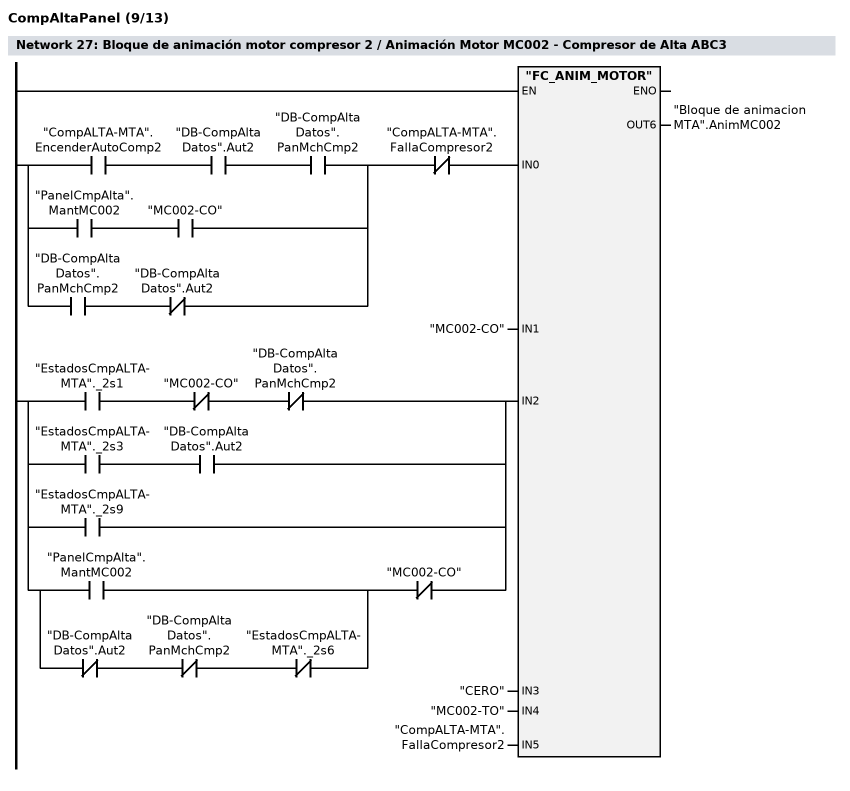
   RUNG wire#powerrail
      "FC_ANIM_MOTOR"(IN0 := wire#w2, IN2 := wire#w4, IN1 := "MC002-CO", IN3 := "CERO", IN4 := "MC002-TO", IN5 := "CompALTA-MTA".FallaCompresor2, OUT6 => "Bloque de animacion MTA".AnimMC002)
   END_RUNG
   RUNG wire#powerrail
      Contact( "CompALTA-MTA".EncenderAutoComp2 )
      Contact( "DB-CompAltaDatos".Aut2 )
      Contact( "DB-CompAltaDatos".PanMchCmp2 )
      wire#w1
      I_Contact( "CompALTA-MTA".FallaCompresor2 )
   END_RUNG wire#w2
   RUNG wire#powerrail
      Contact( "PanelCmpAlta".MantMC002 )
      Contact( "MC002-CO" )
   END_RUNG wire#w1
   RUNG wire#powerrail
      Contact( "DB-CompAltaDatos".PanMchCmp2 )
      I_Contact( "DB-CompAltaDatos".Aut2 )
   END_RUNG wire#w1
   RUNG wire#powerrail
      Contact( "EstadosCmpALTA-MTA"._2s1 )
      I_Contact( "MC002-CO" )
      I_Contact( "DB-CompAltaDatos".PanMchCmp2 )
   END_RUNG wire#w4
   RUNG wire#powerrail
      Contact( "EstadosCmpALTA-MTA"._2s3 )
      Contact( "DB-CompAltaDatos".Aut2 )
   END_RUNG wire#w4
   RUNG wire#powerrail
      Contact( "EstadosCmpALTA-MTA"._2s9 )
   END_RUNG wire#w4
   RUNG wire#powerrail
      Contact( "PanelCmpAlta".MantMC002 )
      wire#w3
      I_Contact( "MC002-CO" )
   END_RUNG wire#w4
   RUNG wire#powerrail
      I_Contact( "DB-CompAltaDatos".Aut2 )
      I_Contact( "DB-CompAltaDatos".PanMchCmp2 )
      I_Contact( "EstadosCmpALTA-MTA"._2s6 )
   END_RUNG wire#w3
   // the same network as SCL:
   "FC_ANIM_MOTOR"(IN0 := (("CompALTA-MTA".EncenderAutoComp2 AND "DB-CompAltaDatos".Aut2 AND "DB-CompAltaDatos".PanMchCmp2) OR ("PanelCmpAlta".MantMC002 AND "MC002-CO") OR ("DB-CompAltaDatos".PanMchCmp2 AND NOT "DB-CompAltaDatos".Aut2)) AND NOT "CompALTA-MTA".FallaCompresor2,
                   IN1 := "MC002-CO",
                   IN2 := ("EstadosCmpALTA-MTA"._2s1 AND NOT "MC002-CO" AND NOT "DB-CompAltaDatos".PanMchCmp2) OR ("EstadosCmpALTA-MTA"._2s3 AND "DB-CompAltaDatos".Aut2) OR "EstadosCmpALTA-MTA"._2s9 OR (("PanelCmpAlta".MantMC002 OR (NOT "DB-CompAltaDatos".Aut2 AND NOT "DB-CompAltaDatos".PanMchCmp2 AND NOT "EstadosCmpALTA-MTA"._2s6)) AND NOT "MC002-CO"),
                   IN3 := "CERO",
                   IN4 := "MC002-TO",
                   IN5 := "CompALTA-MTA".FallaCompresor2,
                   OUT6 => "Bloque de animacion MTA".AnimMC002);
END_REGION

REGION Network 28: Bloque de animación motor compresor 3 / Animación Motor MC003 - Compresor de Alta BELLIS
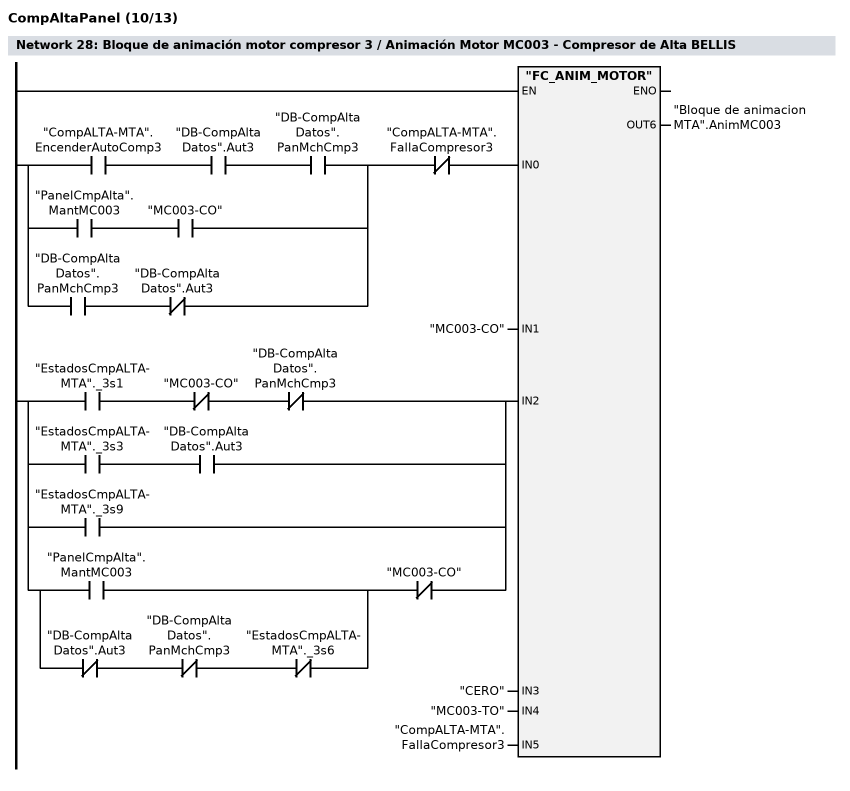
   RUNG wire#powerrail
      "FC_ANIM_MOTOR"(IN0 := wire#w2, IN2 := wire#w4, IN1 := "MC003-CO", IN3 := "CERO", IN4 := "MC003-TO", IN5 := "CompALTA-MTA".FallaCompresor3, OUT6 => "Bloque de animacion MTA".AnimMC003)
   END_RUNG
   RUNG wire#powerrail
      Contact( "CompALTA-MTA".EncenderAutoComp3 )
      Contact( "DB-CompAltaDatos".Aut3 )
      Contact( "DB-CompAltaDatos".PanMchCmp3 )
      wire#w1
      I_Contact( "CompALTA-MTA".FallaCompresor3 )
   END_RUNG wire#w2
   RUNG wire#powerrail
      Contact( "PanelCmpAlta".MantMC003 )
      Contact( "MC003-CO" )
   END_RUNG wire#w1
   RUNG wire#powerrail
      Contact( "DB-CompAltaDatos".PanMchCmp3 )
      I_Contact( "DB-CompAltaDatos".Aut3 )
   END_RUNG wire#w1
   RUNG wire#powerrail
      Contact( "EstadosCmpALTA-MTA"._3s1 )
      I_Contact( "MC003-CO" )
      I_Contact( "DB-CompAltaDatos".PanMchCmp3 )
   END_RUNG wire#w4
   RUNG wire#powerrail
      Contact( "EstadosCmpALTA-MTA"._3s3 )
      Contact( "DB-CompAltaDatos".Aut3 )
   END_RUNG wire#w4
   RUNG wire#powerrail
      Contact( "EstadosCmpALTA-MTA"._3s9 )
   END_RUNG wire#w4
   RUNG wire#powerrail
      Contact( "PanelCmpAlta".MantMC003 )
      wire#w3
      I_Contact( "MC003-CO" )
   END_RUNG wire#w4
   RUNG wire#powerrail
      I_Contact( "DB-CompAltaDatos".Aut3 )
      I_Contact( "DB-CompAltaDatos".PanMchCmp3 )
      I_Contact( "EstadosCmpALTA-MTA"._3s6 )
   END_RUNG wire#w3
   // the same network as SCL:
   "FC_ANIM_MOTOR"(IN0 := (("CompALTA-MTA".EncenderAutoComp3 AND "DB-CompAltaDatos".Aut3 AND "DB-CompAltaDatos".PanMchCmp3) OR ("PanelCmpAlta".MantMC003 AND "MC003-CO") OR ("DB-CompAltaDatos".PanMchCmp3 AND NOT "DB-CompAltaDatos".Aut3)) AND NOT "CompALTA-MTA".FallaCompresor3,
                   IN1 := "MC003-CO",
                   IN2 := ("EstadosCmpALTA-MTA"._3s1 AND NOT "MC003-CO" AND NOT "DB-CompAltaDatos".PanMchCmp3) OR ("EstadosCmpALTA-MTA"._3s3 AND "DB-CompAltaDatos".Aut3) OR "EstadosCmpALTA-MTA"._3s9 OR (("PanelCmpAlta".MantMC003 OR (NOT "DB-CompAltaDatos".Aut3 AND NOT "DB-CompAltaDatos".PanMchCmp3 AND NOT "EstadosCmpALTA-MTA"._3s6)) AND NOT "MC003-CO"),
                   IN3 := "CERO",
                   IN4 := "MC003-TO",
                   IN5 := "CompALTA-MTA".FallaCompresor3,
                   OUT6 => "Bloque de animacion MTA".AnimMC003);
END_REGION

REGION Network 29: Bloque de animación motor compresor 4 / Animación Motor MC004 - Compresor de Alta ABC4
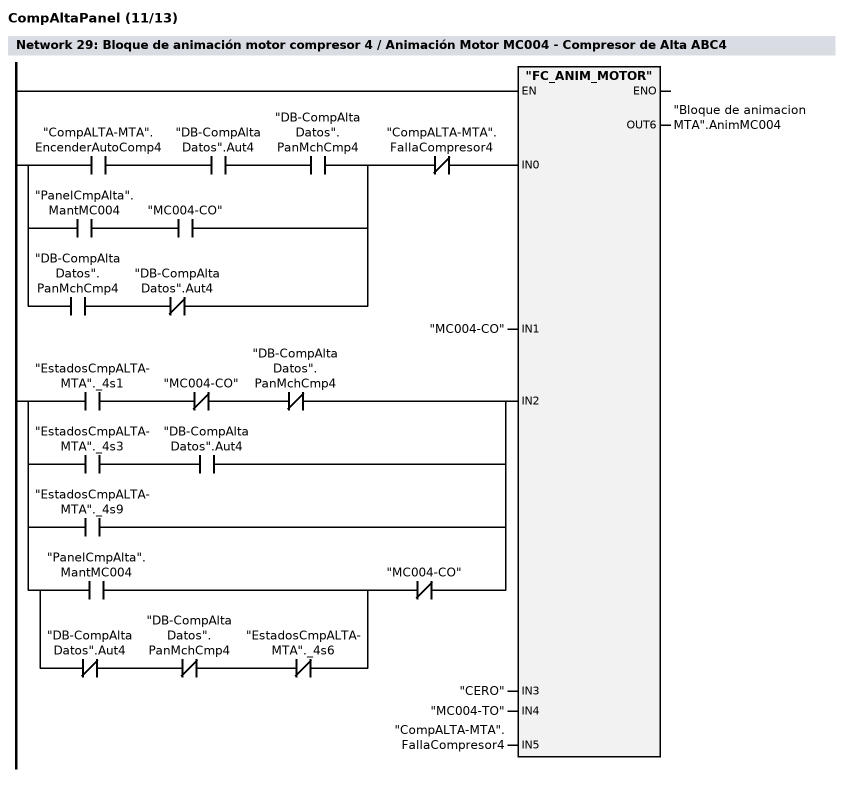
   RUNG wire#powerrail
      "FC_ANIM_MOTOR"(IN0 := wire#w2, IN2 := wire#w4, IN1 := "MC004-CO", IN3 := "CERO", IN4 := "MC004-TO", IN5 := "CompALTA-MTA".FallaCompresor4, OUT6 => "Bloque de animacion MTA".AnimMC004)
   END_RUNG
   RUNG wire#powerrail
      Contact( "CompALTA-MTA".EncenderAutoComp4 )
      Contact( "DB-CompAltaDatos".Aut4 )
      Contact( "DB-CompAltaDatos".PanMchCmp4 )
      wire#w1
      I_Contact( "CompALTA-MTA".FallaCompresor4 )
   END_RUNG wire#w2
   RUNG wire#powerrail
      Contact( "PanelCmpAlta".MantMC004 )
      Contact( "MC004-CO" )
   END_RUNG wire#w1
   RUNG wire#powerrail
      Contact( "DB-CompAltaDatos".PanMchCmp4 )
      I_Contact( "DB-CompAltaDatos".Aut4 )
   END_RUNG wire#w1
   RUNG wire#powerrail
      Contact( "EstadosCmpALTA-MTA"._4s1 )
      I_Contact( "MC004-CO" )
      I_Contact( "DB-CompAltaDatos".PanMchCmp4 )
   END_RUNG wire#w4
   RUNG wire#powerrail
      Contact( "EstadosCmpALTA-MTA"._4s3 )
      Contact( "DB-CompAltaDatos".Aut4 )
   END_RUNG wire#w4
   RUNG wire#powerrail
      Contact( "EstadosCmpALTA-MTA"._4s9 )
   END_RUNG wire#w4
   RUNG wire#powerrail
      Contact( "PanelCmpAlta".MantMC004 )
      wire#w3
      I_Contact( "MC004-CO" )
   END_RUNG wire#w4
   RUNG wire#powerrail
      I_Contact( "DB-CompAltaDatos".Aut4 )
      I_Contact( "DB-CompAltaDatos".PanMchCmp4 )
      I_Contact( "EstadosCmpALTA-MTA"._4s6 )
   END_RUNG wire#w3
   // the same network as SCL:
   "FC_ANIM_MOTOR"(IN0 := (("CompALTA-MTA".EncenderAutoComp4 AND "DB-CompAltaDatos".Aut4 AND "DB-CompAltaDatos".PanMchCmp4) OR ("PanelCmpAlta".MantMC004 AND "MC004-CO") OR ("DB-CompAltaDatos".PanMchCmp4 AND NOT "DB-CompAltaDatos".Aut4)) AND NOT "CompALTA-MTA".FallaCompresor4,
                   IN1 := "MC004-CO",
                   IN2 := ("EstadosCmpALTA-MTA"._4s1 AND NOT "MC004-CO" AND NOT "DB-CompAltaDatos".PanMchCmp4) OR ("EstadosCmpALTA-MTA"._4s3 AND "DB-CompAltaDatos".Aut4) OR "EstadosCmpALTA-MTA"._4s9 OR (("PanelCmpAlta".MantMC004 OR (NOT "DB-CompAltaDatos".Aut4 AND NOT "DB-CompAltaDatos".PanMchCmp4 AND NOT "EstadosCmpALTA-MTA"._4s6)) AND NOT "MC004-CO"),
                   IN3 := "CERO",
                   IN4 := "MC004-TO",
                   IN5 := "CompALTA-MTA".FallaCompresor4,
                   OUT6 => "Bloque de animacion MTA".AnimMC004);
END_REGION

REGION Network 30: Bloque de animación motor compresor 5 / Animación Motor MC005 - Compresor de Alta ABC5
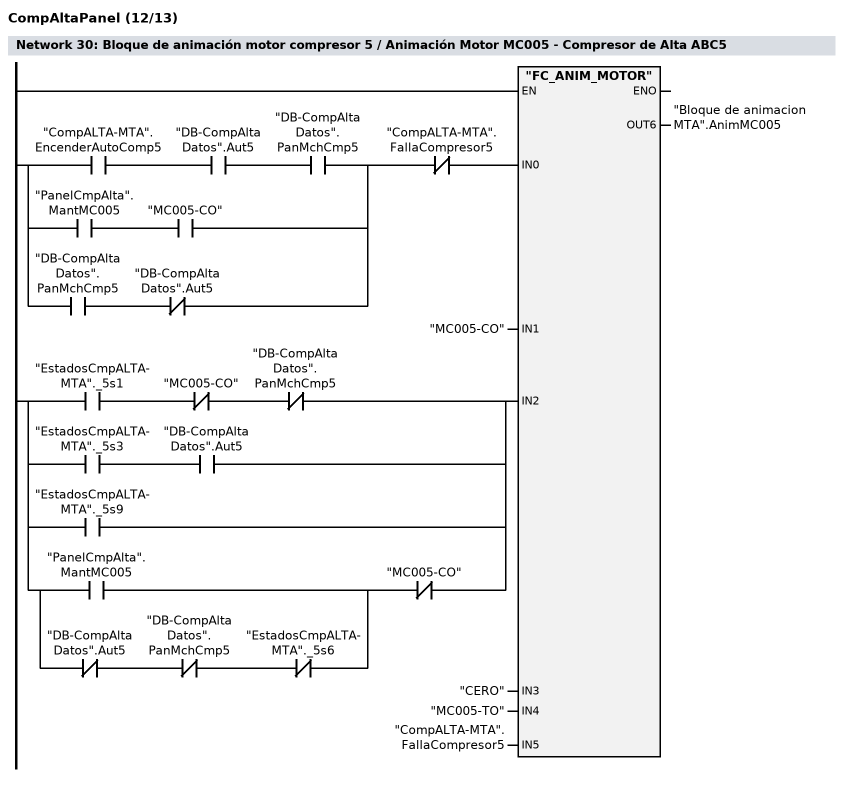
   RUNG wire#powerrail
      "FC_ANIM_MOTOR"(IN0 := wire#w2, IN2 := wire#w4, IN1 := "MC005-CO", IN3 := "CERO", IN4 := "MC005-TO", IN5 := "CompALTA-MTA".FallaCompresor5, OUT6 => "Bloque de animacion MTA".AnimMC005)
   END_RUNG
   RUNG wire#powerrail
      Contact( "CompALTA-MTA".EncenderAutoComp5 )
      Contact( "DB-CompAltaDatos".Aut5 )
      Contact( "DB-CompAltaDatos".PanMchCmp5 )
      wire#w1
      I_Contact( "CompALTA-MTA".FallaCompresor5 )
   END_RUNG wire#w2
   RUNG wire#powerrail
      Contact( "PanelCmpAlta".MantMC005 )
      Contact( "MC005-CO" )
   END_RUNG wire#w1
   RUNG wire#powerrail
      Contact( "DB-CompAltaDatos".PanMchCmp5 )
      I_Contact( "DB-CompAltaDatos".Aut5 )
   END_RUNG wire#w1
   RUNG wire#powerrail
      Contact( "EstadosCmpALTA-MTA"._5s1 )
      I_Contact( "MC005-CO" )
      I_Contact( "DB-CompAltaDatos".PanMchCmp5 )
   END_RUNG wire#w4
   RUNG wire#powerrail
      Contact( "EstadosCmpALTA-MTA"._5s3 )
      Contact( "DB-CompAltaDatos".Aut5 )
   END_RUNG wire#w4
   RUNG wire#powerrail
      Contact( "EstadosCmpALTA-MTA"._5s9 )
   END_RUNG wire#w4
   RUNG wire#powerrail
      Contact( "PanelCmpAlta".MantMC005 )
      wire#w3
      I_Contact( "MC005-CO" )
   END_RUNG wire#w4
   RUNG wire#powerrail
      I_Contact( "DB-CompAltaDatos".Aut5 )
      I_Contact( "DB-CompAltaDatos".PanMchCmp5 )
      I_Contact( "EstadosCmpALTA-MTA"._5s6 )
   END_RUNG wire#w3
   // the same network as SCL:
   "FC_ANIM_MOTOR"(IN0 := (("CompALTA-MTA".EncenderAutoComp5 AND "DB-CompAltaDatos".Aut5 AND "DB-CompAltaDatos".PanMchCmp5) OR ("PanelCmpAlta".MantMC005 AND "MC005-CO") OR ("DB-CompAltaDatos".PanMchCmp5 AND NOT "DB-CompAltaDatos".Aut5)) AND NOT "CompALTA-MTA".FallaCompresor5,
                   IN1 := "MC005-CO",
                   IN2 := ("EstadosCmpALTA-MTA"._5s1 AND NOT "MC005-CO" AND NOT "DB-CompAltaDatos".PanMchCmp5) OR ("EstadosCmpALTA-MTA"._5s3 AND "DB-CompAltaDatos".Aut5) OR "EstadosCmpALTA-MTA"._5s9 OR (("PanelCmpAlta".MantMC005 OR (NOT "DB-CompAltaDatos".Aut5 AND NOT "DB-CompAltaDatos".PanMchCmp5 AND NOT "EstadosCmpALTA-MTA"._5s6)) AND NOT "MC005-CO"),
                   IN3 := "CERO",
                   IN4 := "MC005-TO",
                   IN5 := "CompALTA-MTA".FallaCompresor5,
                   OUT6 => "Bloque de animacion MTA".AnimMC005);
END_REGION

REGION Network 31: Bloque de animación motor compresor 6 / Animación Motor MC005 - Compresor de Alta ABC5
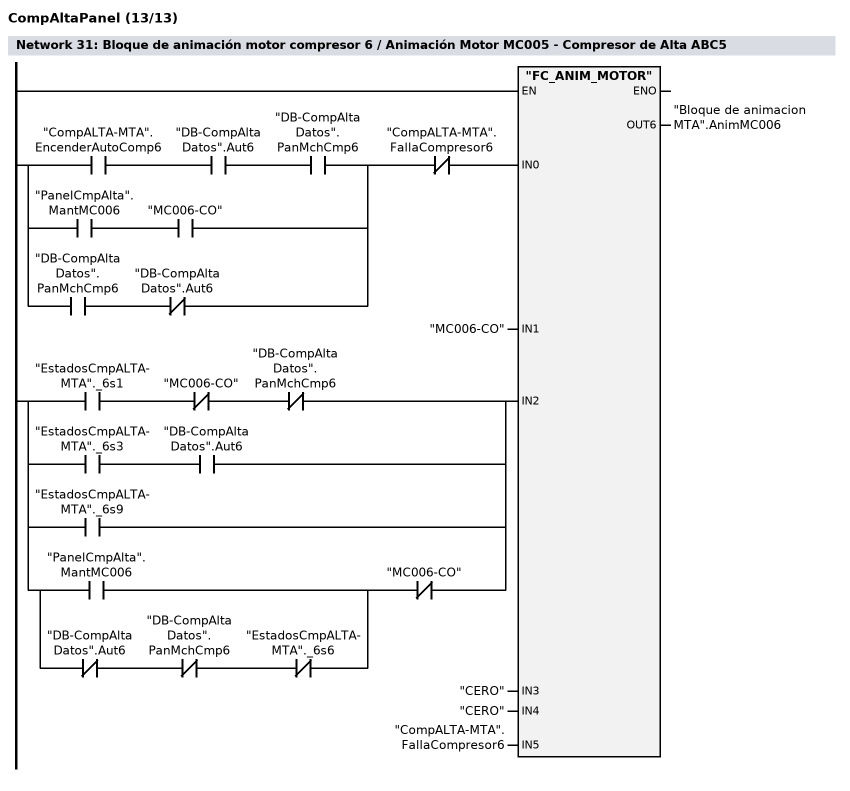
   RUNG wire#powerrail
      "FC_ANIM_MOTOR"(IN0 := wire#w2, IN2 := wire#w4, IN1 := "MC006-CO", IN3 := "CERO", IN4 := "CERO", IN5 := "CompALTA-MTA".FallaCompresor6, OUT6 => "Bloque de animacion MTA".AnimMC006)
   END_RUNG
   RUNG wire#powerrail
      Contact( "CompALTA-MTA".EncenderAutoComp6 )
      Contact( "DB-CompAltaDatos".Aut6 )
      Contact( "DB-CompAltaDatos".PanMchCmp6 )
      wire#w1
      I_Contact( "CompALTA-MTA".FallaCompresor6 )
   END_RUNG wire#w2
   RUNG wire#powerrail
      Contact( "PanelCmpAlta".MantMC006 )
      Contact( "MC006-CO" )
   END_RUNG wire#w1
   RUNG wire#powerrail
      Contact( "DB-CompAltaDatos".PanMchCmp6 )
      I_Contact( "DB-CompAltaDatos".Aut6 )
   END_RUNG wire#w1
   RUNG wire#powerrail
      Contact( "EstadosCmpALTA-MTA"._6s1 )
      I_Contact( "MC006-CO" )
      I_Contact( "DB-CompAltaDatos".PanMchCmp6 )
   END_RUNG wire#w4
   RUNG wire#powerrail
      Contact( "EstadosCmpALTA-MTA"._6s3 )
      Contact( "DB-CompAltaDatos".Aut6 )
   END_RUNG wire#w4
   RUNG wire#powerrail
      Contact( "EstadosCmpALTA-MTA"._6s9 )
   END_RUNG wire#w4
   RUNG wire#powerrail
      Contact( "PanelCmpAlta".MantMC006 )
      wire#w3
      I_Contact( "MC006-CO" )
   END_RUNG wire#w4
   RUNG wire#powerrail
      I_Contact( "DB-CompAltaDatos".Aut6 )
      I_Contact( "DB-CompAltaDatos".PanMchCmp6 )
      I_Contact( "EstadosCmpALTA-MTA"._6s6 )
   END_RUNG wire#w3
   // the same network as SCL:
   "FC_ANIM_MOTOR"(IN0 := (("CompALTA-MTA".EncenderAutoComp6 AND "DB-CompAltaDatos".Aut6 AND "DB-CompAltaDatos".PanMchCmp6) OR ("PanelCmpAlta".MantMC006 AND "MC006-CO") OR ("DB-CompAltaDatos".PanMchCmp6 AND NOT "DB-CompAltaDatos".Aut6)) AND NOT "CompALTA-MTA".FallaCompresor6,
                   IN1 := "MC006-CO",
                   IN2 := ("EstadosCmpALTA-MTA"._6s1 AND NOT "MC006-CO" AND NOT "DB-CompAltaDatos".PanMchCmp6) OR ("EstadosCmpALTA-MTA"._6s3 AND "DB-CompAltaDatos".Aut6) OR "EstadosCmpALTA-MTA"._6s9 OR (("PanelCmpAlta".MantMC006 OR (NOT "DB-CompAltaDatos".Aut6 AND NOT "DB-CompAltaDatos".PanMchCmp6 AND NOT "EstadosCmpALTA-MTA"._6s6)) AND NOT "MC006-CO"),
                   IN3 := "CERO",
                   IN4 := "CERO",
                   IN5 := "CompALTA-MTA".FallaCompresor6,
                   OUT6 => "Bloque de animacion MTA".AnimMC006);
END_REGION
END_FUNCTION

FUNCTION "ModoManualAlta" : Void   // FC48, LAD
{ S7_Optimized_Access := 'FALSE' }
VERSION : 0.1
   VAR_TEMP   // added for the SCL form of the ladder/FBD networks
      _w1 : Bool;
      _s5time1 : S5Time;
   END_VAR
BEGIN

REGION Network 1
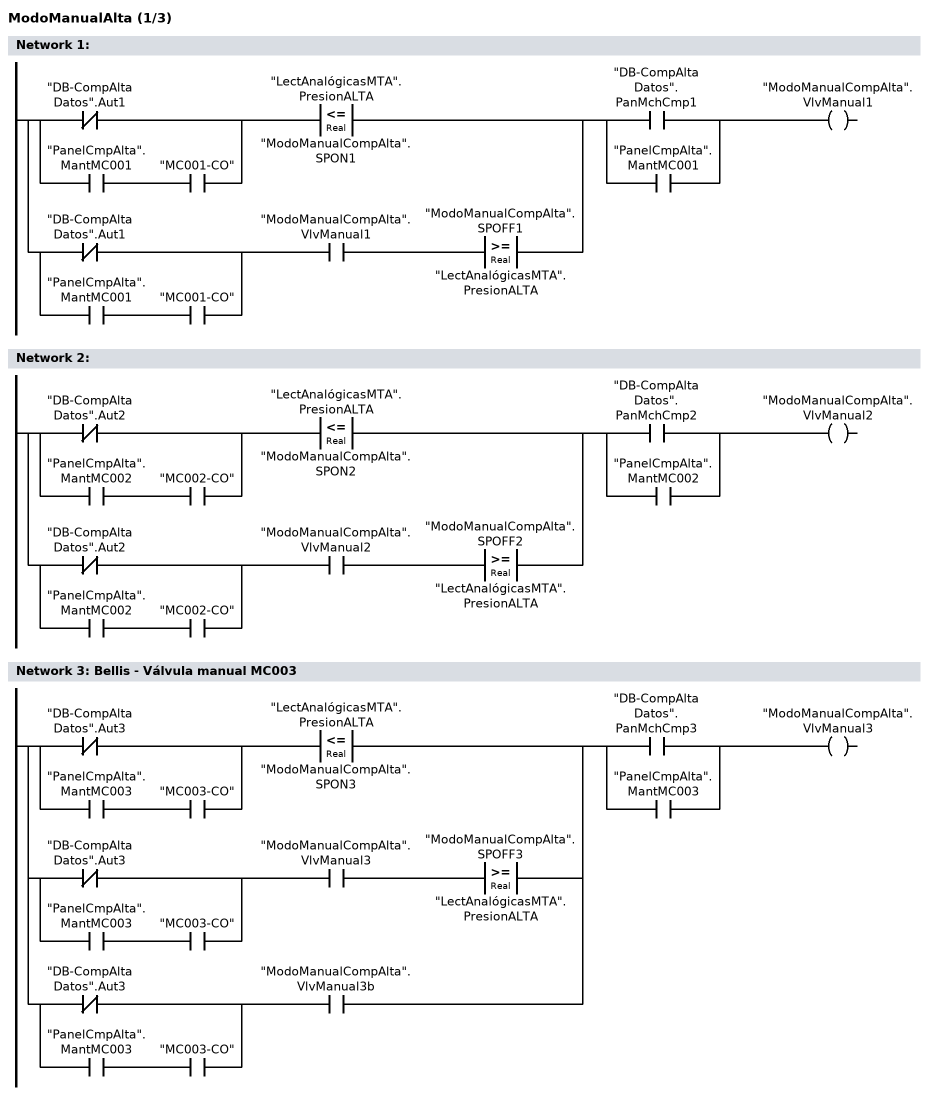
   RUNG wire#powerrail
      I_Contact( "DB-CompAltaDatos".Aut1 )
      wire#w1
      { S7_Templates := "SrcType := Real" } LE_Contact(in1 := "LectAnalógicasMTA".PresionALTA, in2 := "ModoManualCompAlta".SPON1)
      wire#w2
      Contact( "DB-CompAltaDatos".PanMchCmp1 )
      wire#w4
      Coil( "ModoManualCompAlta".VlvManual1 )
   END_RUNG
   RUNG wire#powerrail
      Contact( "PanelCmpAlta".MantMC001 )
      Contact( "MC001-CO" )
   END_RUNG wire#w1
   RUNG wire#powerrail
      I_Contact( "DB-CompAltaDatos".Aut1 )
      wire#w3
      Contact( "ModoManualCompAlta".VlvManual1 )
      { S7_Templates := "SrcType := Real" } GE_Contact(in1 := "ModoManualCompAlta".SPOFF1, in2 := "LectAnalógicasMTA".PresionALTA)
   END_RUNG wire#w2
   RUNG wire#powerrail
      Contact( "PanelCmpAlta".MantMC001 )
      Contact( "MC001-CO" )
   END_RUNG wire#w3
   RUNG wire#w2
      Contact( "PanelCmpAlta".MantMC001 )
   END_RUNG wire#w4
   // the same network as SCL:
   "ModoManualCompAlta".VlvManual1 := (((NOT "DB-CompAltaDatos".Aut1 OR ("PanelCmpAlta".MantMC001 AND "MC001-CO")) AND ("LectAnalógicasMTA".PresionALTA <= "ModoManualCompAlta".SPON1)) OR ((NOT "DB-CompAltaDatos".Aut1 OR ("PanelCmpAlta".MantMC001 AND "MC001-CO")) AND "ModoManualCompAlta".VlvManual1 AND ("ModoManualCompAlta".SPOFF1 >= "LectAnalógicasMTA".PresionALTA))) AND ("DB-CompAltaDatos".PanMchCmp1 OR "PanelCmpAlta".MantMC001);
END_REGION

REGION Network 2
   RUNG wire#powerrail
      I_Contact( "DB-CompAltaDatos".Aut2 )
      wire#w1
      { S7_Templates := "SrcType := Real" } LE_Contact(in1 := "LectAnalógicasMTA".PresionALTA, in2 := "ModoManualCompAlta".SPON2)
      wire#w2
      Contact( "DB-CompAltaDatos".PanMchCmp2 )
      wire#w4
      Coil( "ModoManualCompAlta".VlvManual2 )
   END_RUNG
   RUNG wire#powerrail
      Contact( "PanelCmpAlta".MantMC002 )
      Contact( "MC002-CO" )
   END_RUNG wire#w1
   RUNG wire#powerrail
      I_Contact( "DB-CompAltaDatos".Aut2 )
      wire#w3
      Contact( "ModoManualCompAlta".VlvManual2 )
      { S7_Templates := "SrcType := Real" } GE_Contact(in1 := "ModoManualCompAlta".SPOFF2, in2 := "LectAnalógicasMTA".PresionALTA)
   END_RUNG wire#w2
   RUNG wire#powerrail
      Contact( "PanelCmpAlta".MantMC002 )
      Contact( "MC002-CO" )
   END_RUNG wire#w3
   RUNG wire#w2
      Contact( "PanelCmpAlta".MantMC002 )
   END_RUNG wire#w4
   // the same network as SCL:
   "ModoManualCompAlta".VlvManual2 := (((NOT "DB-CompAltaDatos".Aut2 OR ("PanelCmpAlta".MantMC002 AND "MC002-CO")) AND ("LectAnalógicasMTA".PresionALTA <= "ModoManualCompAlta".SPON2)) OR ((NOT "DB-CompAltaDatos".Aut2 OR ("PanelCmpAlta".MantMC002 AND "MC002-CO")) AND "ModoManualCompAlta".VlvManual2 AND ("ModoManualCompAlta".SPOFF2 >= "LectAnalógicasMTA".PresionALTA))) AND ("DB-CompAltaDatos".PanMchCmp2 OR "PanelCmpAlta".MantMC002);
END_REGION

REGION Network 3: Bellis - Válvula manual MC003
   RUNG wire#powerrail
      I_Contact( "DB-CompAltaDatos".Aut3 )
      wire#w1
      { S7_Templates := "SrcType := Real" } LE_Contact(in1 := "LectAnalógicasMTA".PresionALTA, in2 := "ModoManualCompAlta".SPON3)
      wire#w2
      Contact( "DB-CompAltaDatos".PanMchCmp3 )
      wire#w5
      Coil( "ModoManualCompAlta".VlvManual3 )
   END_RUNG
   RUNG wire#powerrail
      Contact( "PanelCmpAlta".MantMC003 )
      Contact( "MC003-CO" )
   END_RUNG wire#w1
   RUNG wire#powerrail
      I_Contact( "DB-CompAltaDatos".Aut3 )
      wire#w3
      Contact( "ModoManualCompAlta".VlvManual3 )
      { S7_Templates := "SrcType := Real" } GE_Contact(in1 := "ModoManualCompAlta".SPOFF3, in2 := "LectAnalógicasMTA".PresionALTA)
   END_RUNG wire#w2
   RUNG wire#powerrail
      Contact( "PanelCmpAlta".MantMC003 )
      Contact( "MC003-CO" )
   END_RUNG wire#w3
   RUNG wire#powerrail
      I_Contact( "DB-CompAltaDatos".Aut3 )
      wire#w4
      Contact( "ModoManualCompAlta".VlvManual3b )
   END_RUNG wire#w2
   RUNG wire#powerrail
      Contact( "PanelCmpAlta".MantMC003 )
      Contact( "MC003-CO" )
   END_RUNG wire#w4
   RUNG wire#w2
      Contact( "PanelCmpAlta".MantMC003 )
   END_RUNG wire#w5
   // the same network as SCL:
   "ModoManualCompAlta".VlvManual3 := (((NOT "DB-CompAltaDatos".Aut3 OR ("PanelCmpAlta".MantMC003 AND "MC003-CO")) AND ("LectAnalógicasMTA".PresionALTA <= "ModoManualCompAlta".SPON3)) OR ((NOT "DB-CompAltaDatos".Aut3 OR ("PanelCmpAlta".MantMC003 AND "MC003-CO")) AND "ModoManualCompAlta".VlvManual3 AND ("ModoManualCompAlta".SPOFF3 >= "LectAnalógicasMTA".PresionALTA)) OR ((NOT "DB-CompAltaDatos".Aut3 OR ("PanelCmpAlta".MantMC003 AND "MC003-CO")) AND "ModoManualCompAlta".VlvManual3b)) AND ("DB-CompAltaDatos".PanMchCmp3 OR "PanelCmpAlta".MantMC003);
END_REGION

REGION Network 4: Bellis - Válvula manual MC003b
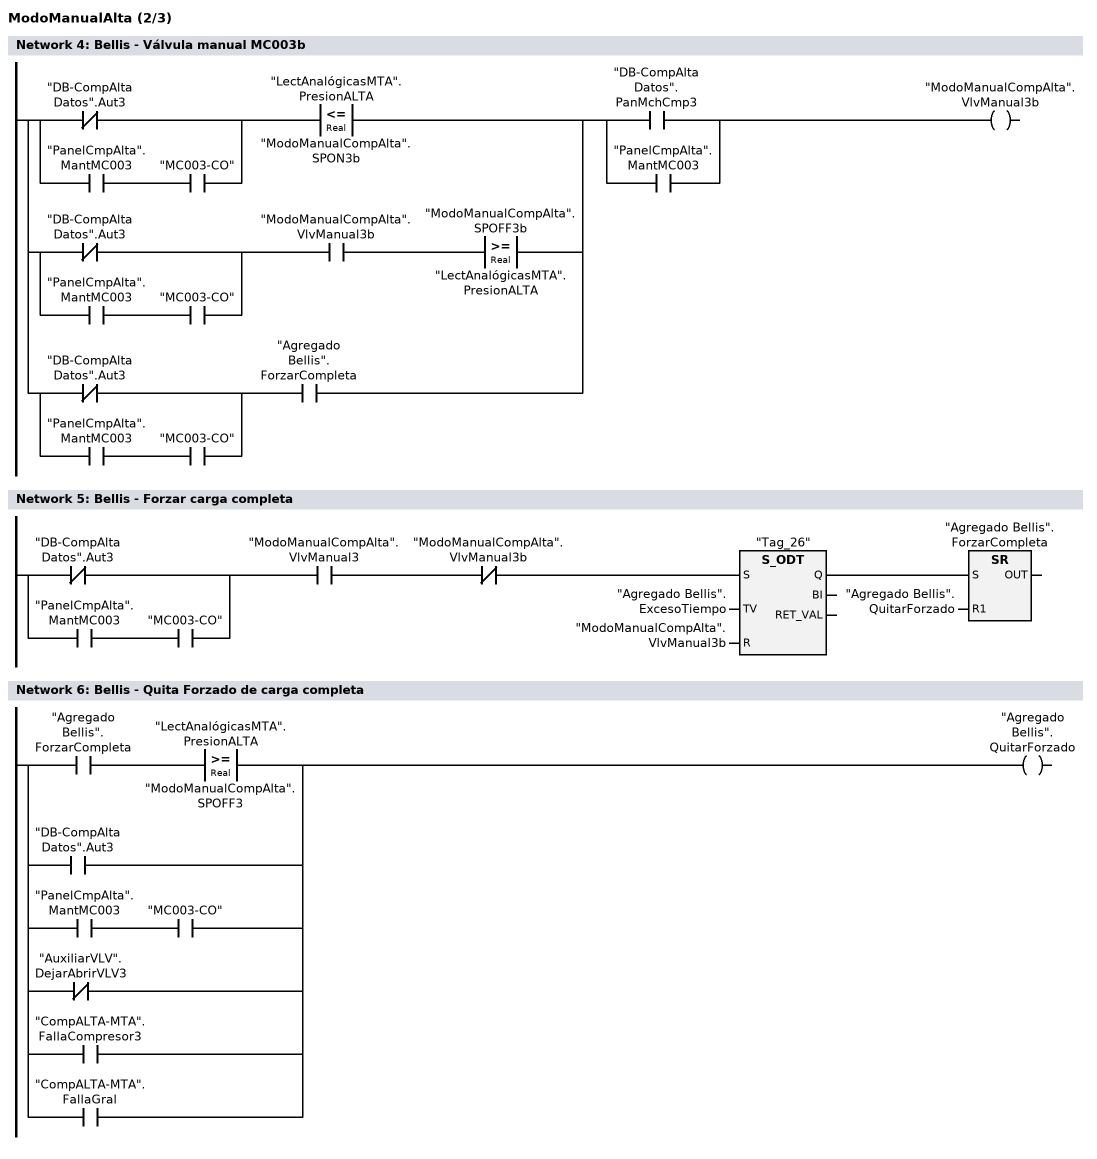
   RUNG wire#powerrail
      I_Contact( "DB-CompAltaDatos".Aut3 )
      wire#w1
      { S7_Templates := "SrcType := Real" } LE_Contact(in1 := "LectAnalógicasMTA".PresionALTA, in2 := "ModoManualCompAlta".SPON3b)
      wire#w2
      Contact( "DB-CompAltaDatos".PanMchCmp3 )
      wire#w5
      Coil( "ModoManualCompAlta".VlvManual3b )
   END_RUNG
   RUNG wire#powerrail
      Contact( "PanelCmpAlta".MantMC003 )
      Contact( "MC003-CO" )
   END_RUNG wire#w1
   RUNG wire#powerrail
      I_Contact( "DB-CompAltaDatos".Aut3 )
      wire#w3
      Contact( "ModoManualCompAlta".VlvManual3b )
      { S7_Templates := "SrcType := Real" } GE_Contact(in1 := "ModoManualCompAlta".SPOFF3b, in2 := "LectAnalógicasMTA".PresionALTA)
   END_RUNG wire#w2
   RUNG wire#powerrail
      Contact( "PanelCmpAlta".MantMC003 )
      Contact( "MC003-CO" )
   END_RUNG wire#w3
   RUNG wire#powerrail
      I_Contact( "DB-CompAltaDatos".Aut3 )
      wire#w4
      Contact( "Agregado Bellis".ForzarCompleta )
   END_RUNG wire#w2
   RUNG wire#powerrail
      Contact( "PanelCmpAlta".MantMC003 )
      Contact( "MC003-CO" )
   END_RUNG wire#w4
   RUNG wire#w2
      Contact( "PanelCmpAlta".MantMC003 )
   END_RUNG wire#w5
   // the same network as SCL:
   "ModoManualCompAlta".VlvManual3b := (((NOT "DB-CompAltaDatos".Aut3 OR ("PanelCmpAlta".MantMC003 AND "MC003-CO")) AND ("LectAnalógicasMTA".PresionALTA <= "ModoManualCompAlta".SPON3b)) OR ((NOT "DB-CompAltaDatos".Aut3 OR ("PanelCmpAlta".MantMC003 AND "MC003-CO")) AND "ModoManualCompAlta".VlvManual3b AND ("ModoManualCompAlta".SPOFF3b >= "LectAnalógicasMTA".PresionALTA)) OR ((NOT "DB-CompAltaDatos".Aut3 OR ("PanelCmpAlta".MantMC003 AND "MC003-CO")) AND "Agregado Bellis".ForzarCompleta)) AND ("DB-CompAltaDatos".PanMchCmp3 OR "PanelCmpAlta".MantMC003);
END_REGION

REGION Network 5: Bellis - Forzar carga completa
   RUNG wire#powerrail
      I_Contact( "DB-CompAltaDatos".Aut3 )
      wire#w1
      Contact( "ModoManualCompAlta".VlvManual3 )
      I_Contact( "ModoManualCompAlta".VlvManual3b )
      S_ODT(T_NO := "Tag_26", TV := "Agregado Bellis".ExcesoTiempo, R := "ModoManualCompAlta".VlvManual3b, BI =>, RET_VAL =>)
      S_SR(operand := "Agregado Bellis".ForzarCompleta, r1 := "Agregado Bellis".QuitarForzado)
   END_RUNG
   RUNG wire#powerrail
      Contact( "PanelCmpAlta".MantMC003 )
      Contact( "MC003-CO" )
   END_RUNG wire#w1
   // the same network as SCL:
   #_s5time1 := S_ODT(T_NO := "Tag_26",
                      S := (NOT "DB-CompAltaDatos".Aut3 OR ("PanelCmpAlta".MantMC003 AND "MC003-CO")) AND "ModoManualCompAlta".VlvManual3 AND NOT "ModoManualCompAlta".VlvManual3b,
                      TV := "Agregado Bellis".ExcesoTiempo,
                      R := "ModoManualCompAlta".VlvManual3b,
                      Q => #_w1);
   IF #_w1 THEN
       "Agregado Bellis".ForzarCompleta := TRUE;   // SR flip-flop
   END_IF;
   IF "Agregado Bellis".QuitarForzado THEN "Agregado Bellis".ForzarCompleta := FALSE; END_IF;
END_REGION

REGION Network 6: Bellis - Quita Forzado de carga completa
   RUNG wire#powerrail
      Contact( "Agregado Bellis".ForzarCompleta )
      { S7_Templates := "SrcType := Real" } GE_Contact(in1 := "LectAnalógicasMTA".PresionALTA, in2 := "ModoManualCompAlta".SPOFF3)
      wire#w1
      Coil( "Agregado Bellis".QuitarForzado )
   END_RUNG
   RUNG wire#powerrail
      Contact( "DB-CompAltaDatos".Aut3 )
   END_RUNG wire#w1
   RUNG wire#powerrail
      Contact( "PanelCmpAlta".MantMC003 )
      Contact( "MC003-CO" )
   END_RUNG wire#w1
   RUNG wire#powerrail
      I_Contact( "AuxiliarVLV".DejarAbrirVLV3 )
   END_RUNG wire#w1
   RUNG wire#powerrail
      Contact( "CompALTA-MTA".FallaCompresor3 )
   END_RUNG wire#w1
   RUNG wire#powerrail
      Contact( "CompALTA-MTA".FallaGral )
   END_RUNG wire#w1
   // the same network as SCL:
   "Agregado Bellis".QuitarForzado := ("Agregado Bellis".ForzarCompleta AND ("LectAnalógicasMTA".PresionALTA >= "ModoManualCompAlta".SPOFF3)) OR "DB-CompAltaDatos".Aut3 OR ("PanelCmpAlta".MantMC003 AND "MC003-CO") OR NOT "AuxiliarVLV".DejarAbrirVLV3 OR "CompALTA-MTA".FallaCompresor3 OR "CompALTA-MTA".FallaGral;
END_REGION

REGION Network 7
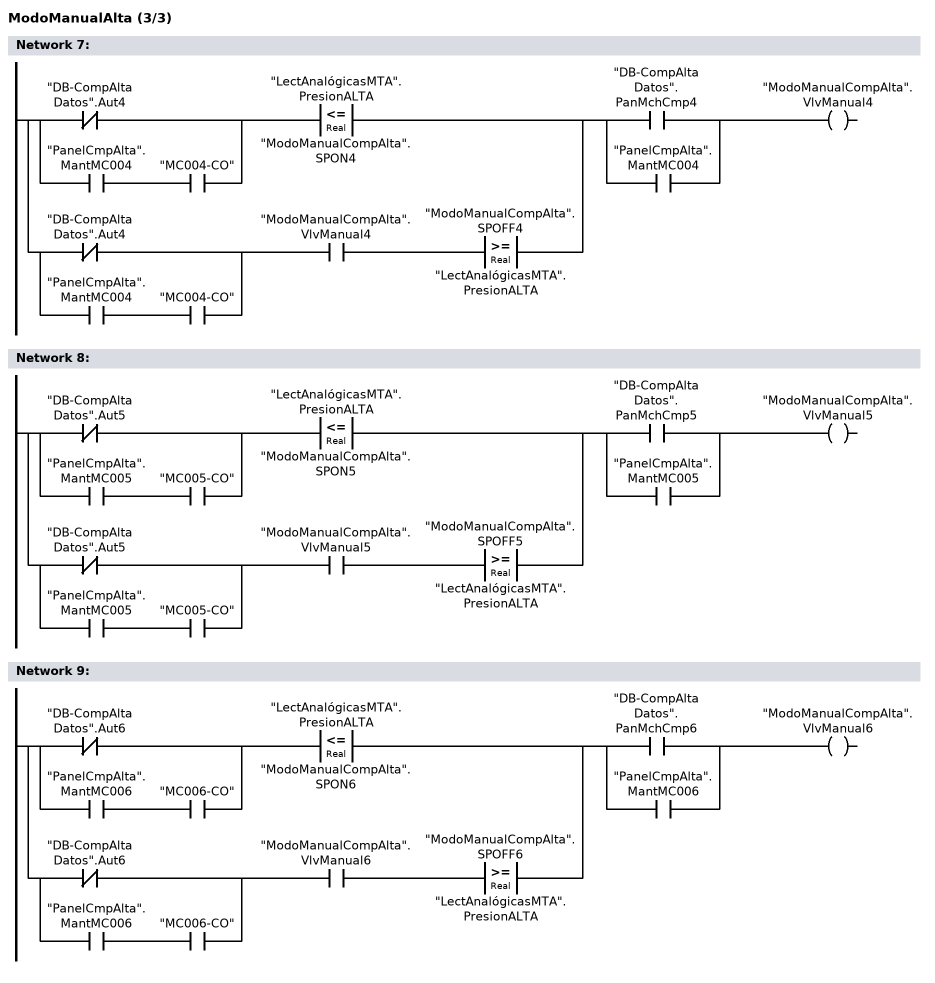
   RUNG wire#powerrail
      I_Contact( "DB-CompAltaDatos".Aut4 )
      wire#w1
      { S7_Templates := "SrcType := Real" } LE_Contact(in1 := "LectAnalógicasMTA".PresionALTA, in2 := "ModoManualCompAlta".SPON4)
      wire#w2
      Contact( "DB-CompAltaDatos".PanMchCmp4 )
      wire#w4
      Coil( "ModoManualCompAlta".VlvManual4 )
   END_RUNG
   RUNG wire#powerrail
      Contact( "PanelCmpAlta".MantMC004 )
      Contact( "MC004-CO" )
   END_RUNG wire#w1
   RUNG wire#powerrail
      I_Contact( "DB-CompAltaDatos".Aut4 )
      wire#w3
      Contact( "ModoManualCompAlta".VlvManual4 )
      { S7_Templates := "SrcType := Real" } GE_Contact(in1 := "ModoManualCompAlta".SPOFF4, in2 := "LectAnalógicasMTA".PresionALTA)
   END_RUNG wire#w2
   RUNG wire#powerrail
      Contact( "PanelCmpAlta".MantMC004 )
      Contact( "MC004-CO" )
   END_RUNG wire#w3
   RUNG wire#w2
      Contact( "PanelCmpAlta".MantMC004 )
   END_RUNG wire#w4
   // the same network as SCL:
   "ModoManualCompAlta".VlvManual4 := (((NOT "DB-CompAltaDatos".Aut4 OR ("PanelCmpAlta".MantMC004 AND "MC004-CO")) AND ("LectAnalógicasMTA".PresionALTA <= "ModoManualCompAlta".SPON4)) OR ((NOT "DB-CompAltaDatos".Aut4 OR ("PanelCmpAlta".MantMC004 AND "MC004-CO")) AND "ModoManualCompAlta".VlvManual4 AND ("ModoManualCompAlta".SPOFF4 >= "LectAnalógicasMTA".PresionALTA))) AND ("DB-CompAltaDatos".PanMchCmp4 OR "PanelCmpAlta".MantMC004);
END_REGION

REGION Network 8
   RUNG wire#powerrail
      I_Contact( "DB-CompAltaDatos".Aut5 )
      wire#w1
      { S7_Templates := "SrcType := Real" } LE_Contact(in1 := "LectAnalógicasMTA".PresionALTA, in2 := "ModoManualCompAlta".SPON5)
      wire#w2
      Contact( "DB-CompAltaDatos".PanMchCmp5 )
      wire#w4
      Coil( "ModoManualCompAlta".VlvManual5 )
   END_RUNG
   RUNG wire#powerrail
      Contact( "PanelCmpAlta".MantMC005 )
      Contact( "MC005-CO" )
   END_RUNG wire#w1
   RUNG wire#powerrail
      I_Contact( "DB-CompAltaDatos".Aut5 )
      wire#w3
      Contact( "ModoManualCompAlta".VlvManual5 )
      { S7_Templates := "SrcType := Real" } GE_Contact(in1 := "ModoManualCompAlta".SPOFF5, in2 := "LectAnalógicasMTA".PresionALTA)
   END_RUNG wire#w2
   RUNG wire#powerrail
      Contact( "PanelCmpAlta".MantMC005 )
      Contact( "MC005-CO" )
   END_RUNG wire#w3
   RUNG wire#w2
      Contact( "PanelCmpAlta".MantMC005 )
   END_RUNG wire#w4
   // the same network as SCL:
   "ModoManualCompAlta".VlvManual5 := (((NOT "DB-CompAltaDatos".Aut5 OR ("PanelCmpAlta".MantMC005 AND "MC005-CO")) AND ("LectAnalógicasMTA".PresionALTA <= "ModoManualCompAlta".SPON5)) OR ((NOT "DB-CompAltaDatos".Aut5 OR ("PanelCmpAlta".MantMC005 AND "MC005-CO")) AND "ModoManualCompAlta".VlvManual5 AND ("ModoManualCompAlta".SPOFF5 >= "LectAnalógicasMTA".PresionALTA))) AND ("DB-CompAltaDatos".PanMchCmp5 OR "PanelCmpAlta".MantMC005);
END_REGION

REGION Network 9
   RUNG wire#powerrail
      I_Contact( "DB-CompAltaDatos".Aut6 )
      wire#w1
      { S7_Templates := "SrcType := Real" } LE_Contact(in1 := "LectAnalógicasMTA".PresionALTA, in2 := "ModoManualCompAlta".SPON6)
      wire#w2
      Contact( "DB-CompAltaDatos".PanMchCmp6 )
      wire#w4
      Coil( "ModoManualCompAlta".VlvManual6 )
   END_RUNG
   RUNG wire#powerrail
      Contact( "PanelCmpAlta".MantMC006 )
      Contact( "MC006-CO" )
   END_RUNG wire#w1
   RUNG wire#powerrail
      I_Contact( "DB-CompAltaDatos".Aut6 )
      wire#w3
      Contact( "ModoManualCompAlta".VlvManual6 )
      { S7_Templates := "SrcType := Real" } GE_Contact(in1 := "ModoManualCompAlta".SPOFF6, in2 := "LectAnalógicasMTA".PresionALTA)
   END_RUNG wire#w2
   RUNG wire#powerrail
      Contact( "PanelCmpAlta".MantMC006 )
      Contact( "MC006-CO" )
   END_RUNG wire#w3
   RUNG wire#w2
      Contact( "PanelCmpAlta".MantMC006 )
   END_RUNG wire#w4
   // the same network as SCL:
   "ModoManualCompAlta".VlvManual6 := (((NOT "DB-CompAltaDatos".Aut6 OR ("PanelCmpAlta".MantMC006 AND "MC006-CO")) AND ("LectAnalógicasMTA".PresionALTA <= "ModoManualCompAlta".SPON6)) OR ((NOT "DB-CompAltaDatos".Aut6 OR ("PanelCmpAlta".MantMC006 AND "MC006-CO")) AND "ModoManualCompAlta".VlvManual6 AND ("ModoManualCompAlta".SPOFF6 >= "LectAnalógicasMTA".PresionALTA))) AND ("DB-CompAltaDatos".PanMchCmp6 OR "PanelCmpAlta".MantMC006);
END_REGION
END_FUNCTION

FUNCTION "PurgaComAlta" : Void   // FC51, LAD
{ S7_Optimized_Access := 'FALSE' }
VERSION : 0.1
// Control de electrovalvulas para realizar purga de compresores, evitando simultaneidad. Con habilitación y seteos de tiempos desde panel.
   VAR_TEMP
      Aux1_MC003 : Word;
      Aux2_MC003 : Word;
      Aux1_MC001 : Word;
      Aux2_MC001 : Word;
      Aux1_MC002 : Word;
      Aux2_MC002 : Word;
      Aux1_MC004 : Word;
      Aux2_MC004 : Word;
      Aux1_MC005 : Word;
      Aux2_MC005 : Word;
      Aux1_MC006 : Word;
      Aux2_MC006 : Word;
   END_VAR
   VAR_TEMP   // added for the SCL form of the ladder/FBD networks
      _w1 : Bool;
      _s5time1 : S5Time;
      _s5time2 : S5Time;
   END_VAR
BEGIN

REGION Network 1
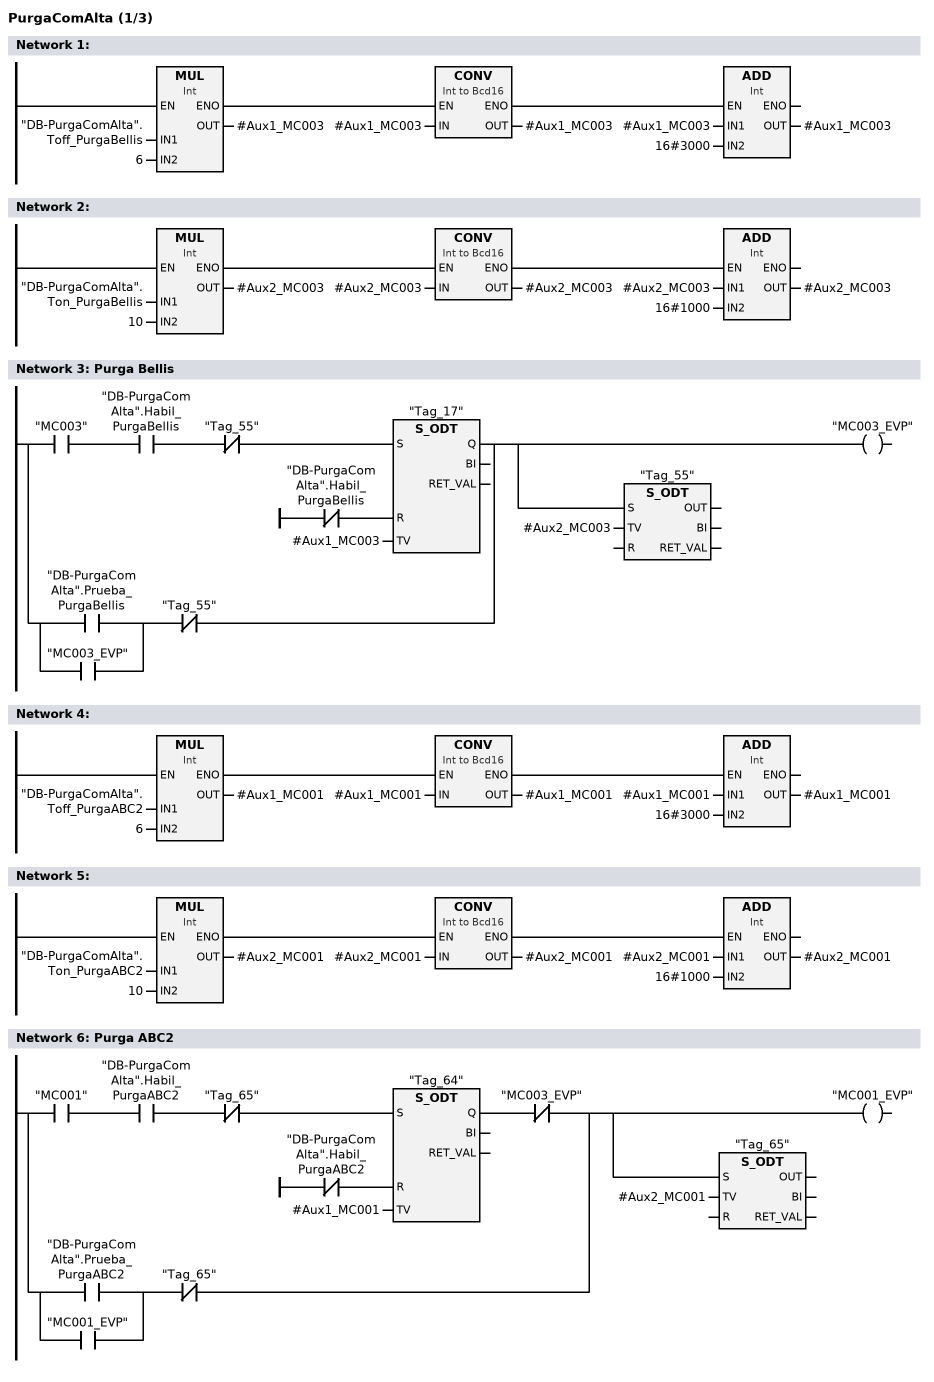
   RUNG wire#powerrail
      { S7_Templates := "SrcType := Int"; S7_GenerateENO := "TRUE" } Mul(in1 := "DB-PurgaComAlta".Toff_PurgaBellis, in2 := 6, out => #Aux1_MC003)
      { S7_Templates := "[SrcType := Int, DestType := Bcd16]"; S7_GenerateENO := "TRUE" } Convert(in := #Aux1_MC003, out => #Aux1_MC003)
      { S7_Templates := "SrcType := Int"; S7_GenerateENO := "TRUE" } Add(in1 := #Aux1_MC003, in2 := 16#3000, out => #Aux1_MC003)
   END_RUNG
   // the same network as SCL:
   // ENO of a box is taken as its EN; it also drops when the box reports an error
   #Aux1_MC003 := "DB-PurgaComAlta".Toff_PurgaBellis * 6;
   #Aux1_MC003 := INT_TO_BCD16(#Aux1_MC003);
   #Aux1_MC003 := #Aux1_MC003 + 16#3000;
END_REGION

REGION Network 2
   RUNG wire#powerrail
      { S7_Templates := "SrcType := Int"; S7_GenerateENO := "TRUE" } Mul(in1 := "DB-PurgaComAlta".Ton_PurgaBellis, in2 := 10, out => #Aux2_MC003)
      { S7_Templates := "[SrcType := Int, DestType := Bcd16]"; S7_GenerateENO := "TRUE" } Convert(in := #Aux2_MC003, out => #Aux2_MC003)
      { S7_Templates := "SrcType := Int"; S7_GenerateENO := "TRUE" } Add(in1 := #Aux2_MC003, in2 := 16#1000, out => #Aux2_MC003)
   END_RUNG
   // the same network as SCL:
   // ENO of a box is taken as its EN; it also drops when the box reports an error
   #Aux2_MC003 := "DB-PurgaComAlta".Ton_PurgaBellis * 10;
   #Aux2_MC003 := INT_TO_BCD16(#Aux2_MC003);
   #Aux2_MC003 := #Aux2_MC003 + 16#1000;
END_REGION
